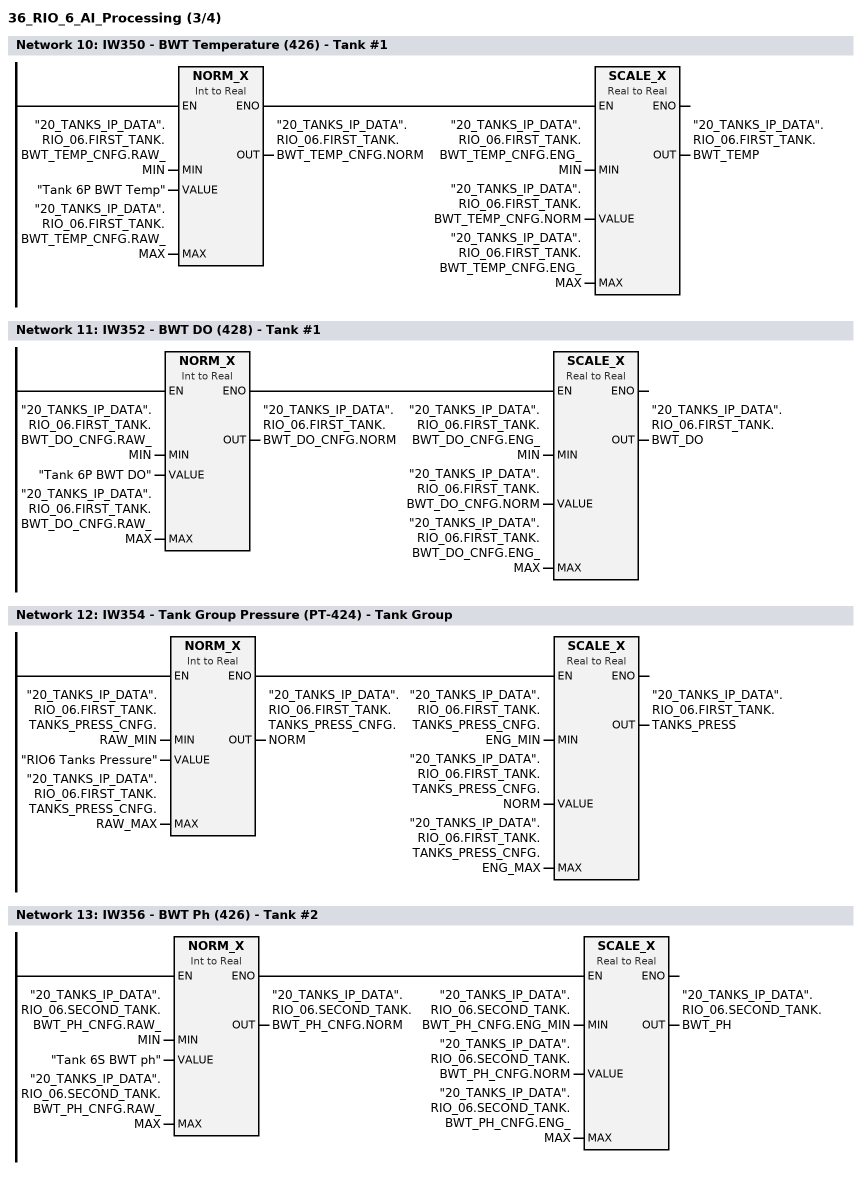
   RUNG wire#powerrail
      { S7_Templates := "[SrcType := Int, DestType := Real]" } Normalize(min := "20_TANKS_IP_DATA".RIO_06.FIRST_TANK.BWT_TEMP_CNFG.RAW_MIN, value := "Tank 6P BWT Temp", max := "20_TANKS_IP_DATA".RIO_06.FIRST_TANK.BWT_TEMP_CNFG.RAW_MAX, out => "20_TANKS_IP_DATA".RIO_06.FIRST_TANK.BWT_TEMP_CNFG.NORM)
      { S7_Templates := "[SrcType := Real, DestType := Real]" } Scale(min := "20_TANKS_IP_DATA".RIO_06.FIRST_TANK.BWT_TEMP_CNFG.ENG_MIN, value := "20_TANKS_IP_DATA".RIO_06.FIRST_TANK.BWT_TEMP_CNFG.NORM, max := "20_TANKS_IP_DATA".RIO_06.FIRST_TANK.BWT_TEMP_CNFG.ENG_MAX, out => "20_TANKS_IP_DATA".RIO_06.FIRST_TANK.BWT_TEMP)
   END_RUNG
   // the same network as SCL:
   "20_TANKS_IP_DATA".RIO_06.FIRST_TANK.BWT_TEMP_CNFG.NORM := NORM_X(MIN := "20_TANKS_IP_DATA".RIO_06.FIRST_TANK.BWT_TEMP_CNFG.RAW_MIN, VALUE := "Tank 6P BWT Temp", MAX := "20_TANKS_IP_DATA".RIO_06.FIRST_TANK.BWT_TEMP_CNFG.RAW_MAX);
   "20_TANKS_IP_DATA".RIO_06.FIRST_TANK.BWT_TEMP := SCALE_X(MIN := "20_TANKS_IP_DATA".RIO_06.FIRST_TANK.BWT_TEMP_CNFG.ENG_MIN, VALUE := "20_TANKS_IP_DATA".RIO_06.FIRST_TANK.BWT_TEMP_CNFG.NORM, MAX := "20_TANKS_IP_DATA".RIO_06.FIRST_TANK.BWT_TEMP_CNFG.ENG_MAX);
END_REGION

REGION Network 11: IW352 - BWT DO (428) - Tank #1
   RUNG wire#powerrail
      { S7_Templates := "[SrcType := Int, DestType := Real]" } Normalize(min := "20_TANKS_IP_DATA".RIO_06.FIRST_TANK.BWT_DO_CNFG.RAW_MIN, value := "Tank 6P BWT DO", max := "20_TANKS_IP_DATA".RIO_06.FIRST_TANK.BWT_DO_CNFG.RAW_MAX, out => "20_TANKS_IP_DATA".RIO_06.FIRST_TANK.BWT_DO_CNFG.NORM)
      { S7_Templates := "[SrcType := Real, DestType := Real]" } Scale(min := "20_TANKS_IP_DATA".RIO_06.FIRST_TANK.BWT_DO_CNFG.ENG_MIN, value := "20_TANKS_IP_DATA".RIO_06.FIRST_TANK.BWT_DO_CNFG.NORM, max := "20_TANKS_IP_DATA".RIO_06.FIRST_TANK.BWT_DO_CNFG.ENG_MAX, out => "20_TANKS_IP_DATA".RIO_06.FIRST_TANK.BWT_DO)
   END_RUNG
   // the same network as SCL:
   "20_TANKS_IP_DATA".RIO_06.FIRST_TANK.BWT_DO_CNFG.NORM := NORM_X(MIN := "20_TANKS_IP_DATA".RIO_06.FIRST_TANK.BWT_DO_CNFG.RAW_MIN, VALUE := "Tank 6P BWT DO", MAX := "20_TANKS_IP_DATA".RIO_06.FIRST_TANK.BWT_DO_CNFG.RAW_MAX);
   "20_TANKS_IP_DATA".RIO_06.FIRST_TANK.BWT_DO := SCALE_X(MIN := "20_TANKS_IP_DATA".RIO_06.FIRST_TANK.BWT_DO_CNFG.ENG_MIN, VALUE := "20_TANKS_IP_DATA".RIO_06.FIRST_TANK.BWT_DO_CNFG.NORM, MAX := "20_TANKS_IP_DATA".RIO_06.FIRST_TANK.BWT_DO_CNFG.ENG_MAX);
END_REGION

REGION Network 12: IW354 - Tank Group Pressure (PT-424) - Tank Group
   RUNG wire#powerrail
      { S7_Templates := "[SrcType := Int, DestType := Real]" } Normalize(min := "20_TANKS_IP_DATA".RIO_06.FIRST_TANK.TANKS_PRESS_CNFG.RAW_MIN, value := "RIO6 Tanks Pressure", max := "20_TANKS_IP_DATA".RIO_06.FIRST_TANK.TANKS_PRESS_CNFG.RAW_MAX, out => "20_TANKS_IP_DATA".RIO_06.FIRST_TANK.TANKS_PRESS_CNFG.NORM)
      { S7_Templates := "[SrcType := Real, DestType := Real]" } Scale(min := "20_TANKS_IP_DATA".RIO_06.FIRST_TANK.TANKS_PRESS_CNFG.ENG_MIN, value := "20_TANKS_IP_DATA".RIO_06.FIRST_TANK.TANKS_PRESS_CNFG.NORM, max := "20_TANKS_IP_DATA".RIO_06.FIRST_TANK.TANKS_PRESS_CNFG.ENG_MAX, out => "20_TANKS_IP_DATA".RIO_06.FIRST_TANK.TANKS_PRESS)
   END_RUNG
   // the same network as SCL:
   "20_TANKS_IP_DATA".RIO_06.FIRST_TANK.TANKS_PRESS_CNFG.NORM := NORM_X(MIN := "20_TANKS_IP_DATA".RIO_06.FIRST_TANK.TANKS_PRESS_CNFG.RAW_MIN, VALUE := "RIO6 Tanks Pressure", MAX := "20_TANKS_IP_DATA".RIO_06.FIRST_TANK.TANKS_PRESS_CNFG.RAW_MAX);
   "20_TANKS_IP_DATA".RIO_06.FIRST_TANK.TANKS_PRESS := SCALE_X(MIN := "20_TANKS_IP_DATA".RIO_06.FIRST_TANK.TANKS_PRESS_CNFG.ENG_MIN, VALUE := "20_TANKS_IP_DATA".RIO_06.FIRST_TANK.TANKS_PRESS_CNFG.NORM, MAX := "20_TANKS_IP_DATA".RIO_06.FIRST_TANK.TANKS_PRESS_CNFG.ENG_MAX);
END_REGION

REGION Network 13: IW356 - BWT Ph (426) - Tank #2
   RUNG wire#powerrail
      { S7_Templates := "[SrcType := Int, DestType := Real]" } Normalize(min := "20_TANKS_IP_DATA".RIO_06.SECOND_TANK.BWT_PH_CNFG.RAW_MIN, value := "Tank 6S BWT ph", max := "20_TANKS_IP_DATA".RIO_06.SECOND_TANK.BWT_PH_CNFG.RAW_MAX, out => "20_TANKS_IP_DATA".RIO_06.SECOND_TANK.BWT_PH_CNFG.NORM)
      { S7_Templates := "[SrcType := Real, DestType := Real]" } Scale(min := "20_TANKS_IP_DATA".RIO_06.SECOND_TANK.BWT_PH_CNFG.ENG_MIN, value := "20_TANKS_IP_DATA".RIO_06.SECOND_TANK.BWT_PH_CNFG.NORM, max := "20_TANKS_IP_DATA".RIO_06.SECOND_TANK.BWT_PH_CNFG.ENG_MAX, out => "20_TANKS_IP_DATA".RIO_06.SECOND_TANK.BWT_PH)
   END_RUNG
   // the same network as SCL:
   "20_TANKS_IP_DATA".RIO_06.SECOND_TANK.BWT_PH_CNFG.NORM := NORM_X(MIN := "20_TANKS_IP_DATA".RIO_06.SECOND_TANK.BWT_PH_CNFG.RAW_MIN, VALUE := "Tank 6S BWT ph", MAX := "20_TANKS_IP_DATA".RIO_06.SECOND_TANK.BWT_PH_CNFG.RAW_MAX);
   "20_TANKS_IP_DATA".RIO_06.SECOND_TANK.BWT_PH := SCALE_X(MIN := "20_TANKS_IP_DATA".RIO_06.SECOND_TANK.BWT_PH_CNFG.ENG_MIN, VALUE := "20_TANKS_IP_DATA".RIO_06.SECOND_TANK.BWT_PH_CNFG.NORM, MAX := "20_TANKS_IP_DATA".RIO_06.SECOND_TANK.BWT_PH_CNFG.ENG_MAX);
END_REGION

REGION Network 14: IW358 - BWT Temperature (426) - Tank #2
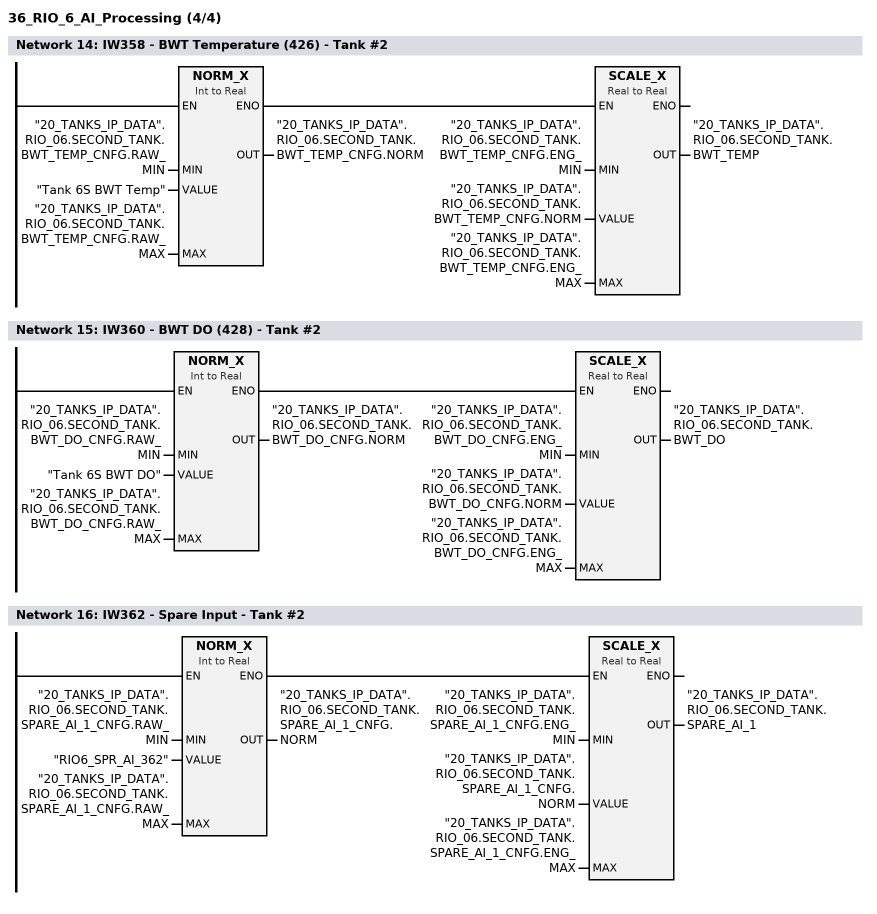
   RUNG wire#powerrail
      { S7_Templates := "[SrcType := Int, DestType := Real]" } Normalize(min := "20_TANKS_IP_DATA".RIO_06.SECOND_TANK.BWT_TEMP_CNFG.RAW_MIN, value := "Tank 6S BWT Temp", max := "20_TANKS_IP_DATA".RIO_06.SECOND_TANK.BWT_TEMP_CNFG.RAW_MAX, out => "20_TANKS_IP_DATA".RIO_06.SECOND_TANK.BWT_TEMP_CNFG.NORM)
      { S7_Templates := "[SrcType := Real, DestType := Real]" } Scale(min := "20_TANKS_IP_DATA".RIO_06.SECOND_TANK.BWT_TEMP_CNFG.ENG_MIN, value := "20_TANKS_IP_DATA".RIO_06.SECOND_TANK.BWT_TEMP_CNFG.NORM, max := "20_TANKS_IP_DATA".RIO_06.SECOND_TANK.BWT_TEMP_CNFG.ENG_MAX, out => "20_TANKS_IP_DATA".RIO_06.SECOND_TANK.BWT_TEMP)
   END_RUNG
   // the same network as SCL:
   "20_TANKS_IP_DATA".RIO_06.SECOND_TANK.BWT_TEMP_CNFG.NORM := NORM_X(MIN := "20_TANKS_IP_DATA".RIO_06.SECOND_TANK.BWT_TEMP_CNFG.RAW_MIN, VALUE := "Tank 6S BWT Temp", MAX := "20_TANKS_IP_DATA".RIO_06.SECOND_TANK.BWT_TEMP_CNFG.RAW_MAX);
   "20_TANKS_IP_DATA".RIO_06.SECOND_TANK.BWT_TEMP := SCALE_X(MIN := "20_TANKS_IP_DATA".RIO_06.SECOND_TANK.BWT_TEMP_CNFG.ENG_MIN, VALUE := "20_TANKS_IP_DATA".RIO_06.SECOND_TANK.BWT_TEMP_CNFG.NORM, MAX := "20_TANKS_IP_DATA".RIO_06.SECOND_TANK.BWT_TEMP_CNFG.ENG_MAX);
END_REGION

REGION Network 15: IW360 - BWT DO (428) - Tank #2
   RUNG wire#powerrail
      { S7_Templates := "[SrcType := Int, DestType := Real]" } Normalize(min := "20_TANKS_IP_DATA".RIO_06.SECOND_TANK.BWT_DO_CNFG.RAW_MIN, value := "Tank 6S BWT DO", max := "20_TANKS_IP_DATA".RIO_06.SECOND_TANK.BWT_DO_CNFG.RAW_MAX, out => "20_TANKS_IP_DATA".RIO_06.SECOND_TANK.BWT_DO_CNFG.NORM)
      { S7_Templates := "[SrcType := Real, DestType := Real]" } Scale(min := "20_TANKS_IP_DATA".RIO_06.SECOND_TANK.BWT_DO_CNFG.ENG_MIN, value := "20_TANKS_IP_DATA".RIO_06.SECOND_TANK.BWT_DO_CNFG.NORM, max := "20_TANKS_IP_DATA".RIO_06.SECOND_TANK.BWT_DO_CNFG.ENG_MAX, out => "20_TANKS_IP_DATA".RIO_06.SECOND_TANK.BWT_DO)
   END_RUNG
   // the same network as SCL:
   "20_TANKS_IP_DATA".RIO_06.SECOND_TANK.BWT_DO_CNFG.NORM := NORM_X(MIN := "20_TANKS_IP_DATA".RIO_06.SECOND_TANK.BWT_DO_CNFG.RAW_MIN, VALUE := "Tank 6S BWT DO", MAX := "20_TANKS_IP_DATA".RIO_06.SECOND_TANK.BWT_DO_CNFG.RAW_MAX);
   "20_TANKS_IP_DATA".RIO_06.SECOND_TANK.BWT_DO := SCALE_X(MIN := "20_TANKS_IP_DATA".RIO_06.SECOND_TANK.BWT_DO_CNFG.ENG_MIN, VALUE := "20_TANKS_IP_DATA".RIO_06.SECOND_TANK.BWT_DO_CNFG.NORM, MAX := "20_TANKS_IP_DATA".RIO_06.SECOND_TANK.BWT_DO_CNFG.ENG_MAX);
END_REGION

REGION Network 16: IW362 - Spare Input - Tank #2
   RUNG wire#powerrail
      { S7_Templates := "[SrcType := Int, DestType := Real]" } Normalize(min := "20_TANKS_IP_DATA".RIO_06.SECOND_TANK.SPARE_AI_1_CNFG.RAW_MIN, value := "RIO6_SPR_AI_362", max := "20_TANKS_IP_DATA".RIO_06.SECOND_TANK.SPARE_AI_1_CNFG.RAW_MAX, out => "20_TANKS_IP_DATA".RIO_06.SECOND_TANK.SPARE_AI_1_CNFG.NORM)
      { S7_Templates := "[SrcType := Real, DestType := Real]" } Scale(min := "20_TANKS_IP_DATA".RIO_06.SECOND_TANK.SPARE_AI_1_CNFG.ENG_MIN, value := "20_TANKS_IP_DATA".RIO_06.SECOND_TANK.SPARE_AI_1_CNFG.NORM, max := "20_TANKS_IP_DATA".RIO_06.SECOND_TANK.SPARE_AI_1_CNFG.ENG_MAX, out => "20_TANKS_IP_DATA".RIO_06.SECOND_TANK.SPARE_AI_1)
   END_RUNG
   // the same network as SCL:
   "20_TANKS_IP_DATA".RIO_06.SECOND_TANK.SPARE_AI_1_CNFG.NORM := NORM_X(MIN := "20_TANKS_IP_DATA".RIO_06.SECOND_TANK.SPARE_AI_1_CNFG.RAW_MIN, VALUE := "RIO6_SPR_AI_362", MAX := "20_TANKS_IP_DATA".RIO_06.SECOND_TANK.SPARE_AI_1_CNFG.RAW_MAX);
   "20_TANKS_IP_DATA".RIO_06.SECOND_TANK.SPARE_AI_1 := SCALE_X(MIN := "20_TANKS_IP_DATA".RIO_06.SECOND_TANK.SPARE_AI_1_CNFG.ENG_MIN, VALUE := "20_TANKS_IP_DATA".RIO_06.SECOND_TANK.SPARE_AI_1_CNFG.NORM, MAX := "20_TANKS_IP_DATA".RIO_06.SECOND_TANK.SPARE_AI_1_CNFG.ENG_MAX);
END_REGION
END_FUNCTION

FUNCTION "37_RIO_7_AI_Processing" : Void   // FC37, LAD
TITLE = Analogue Input Processing (Tank 1 = APT)
{ S7_Optimized_Access := 'TRUE' }
AUTHOR : JRS
VERSION : 0.1
// To process raw inputs prior to code use
BEGIN

REGION Network 1: IW400 - USD Flow (FIT-418) - Tank #1
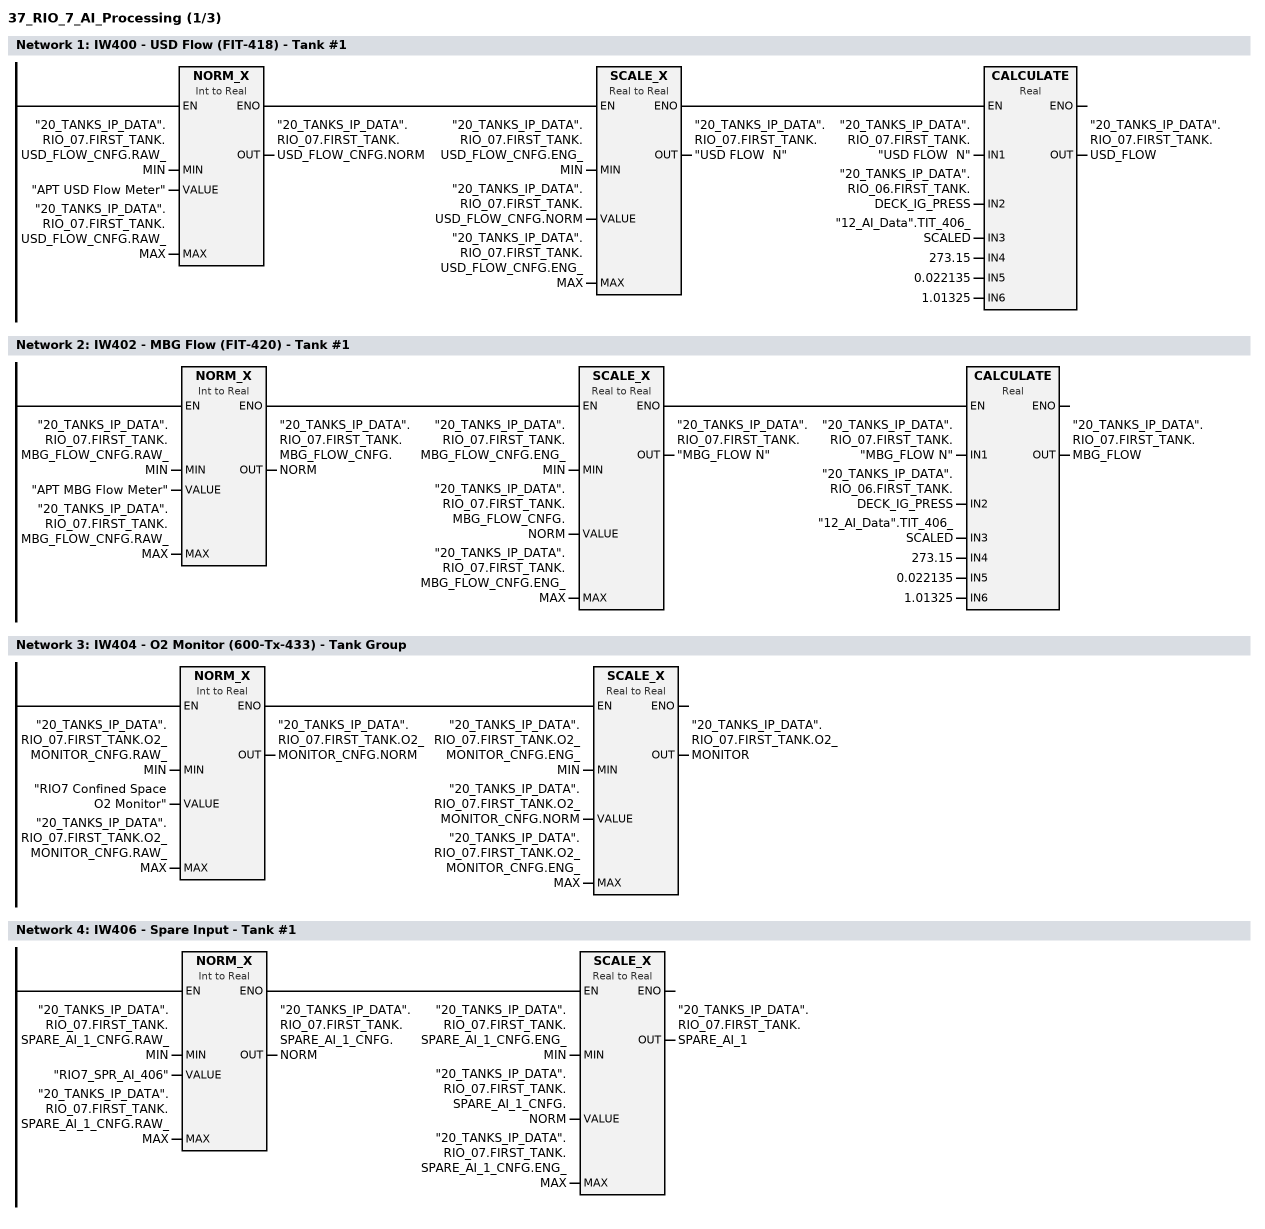
   RUNG wire#powerrail
      { S7_Templates := "[SrcType := Int, DestType := Real]" } Normalize(min := "20_TANKS_IP_DATA".RIO_07.FIRST_TANK.USD_FLOW_CNFG.RAW_MIN, value := "APT USD Flow Meter", max := "20_TANKS_IP_DATA".RIO_07.FIRST_TANK.USD_FLOW_CNFG.RAW_MAX, out => "20_TANKS_IP_DATA".RIO_07.FIRST_TANK.USD_FLOW_CNFG.NORM)
      { S7_Templates := "[SrcType := Real, DestType := Real]" } Scale(min := "20_TANKS_IP_DATA".RIO_07.FIRST_TANK.USD_FLOW_CNFG.ENG_MIN, value := "20_TANKS_IP_DATA".RIO_07.FIRST_TANK.USD_FLOW_CNFG.NORM, max := "20_TANKS_IP_DATA".RIO_07.FIRST_TANK.USD_FLOW_CNFG.ENG_MAX, out => "20_TANKS_IP_DATA".RIO_07.FIRST_TANK."USD FLOW  N")
      { S7_Templates := "SrcType := Real"; S7_Expression := "IN1*(IN2+IN6)/IN6*IN4/(IN3+IN4)" } Calculate(in1 := "20_TANKS_IP_DATA".RIO_07.FIRST_TANK."USD FLOW  N", in2 := "20_TANKS_IP_DATA".RIO_06.FIRST_TANK.DECK_IG_PRESS, in3 := "12_AI_Data".TIT_406_SCALED, in4 := 273.15, in5 := 0.022135, in6 := 1.01325, out => "20_TANKS_IP_DATA".RIO_07.FIRST_TANK.USD_FLOW)
   END_RUNG
   // the same network as SCL:
   "20_TANKS_IP_DATA".RIO_07.FIRST_TANK.USD_FLOW_CNFG.NORM := NORM_X(MIN := "20_TANKS_IP_DATA".RIO_07.FIRST_TANK.USD_FLOW_CNFG.RAW_MIN, VALUE := "APT USD Flow Meter", MAX := "20_TANKS_IP_DATA".RIO_07.FIRST_TANK.USD_FLOW_CNFG.RAW_MAX);
   "20_TANKS_IP_DATA".RIO_07.FIRST_TANK."USD FLOW  N" := SCALE_X(MIN := "20_TANKS_IP_DATA".RIO_07.FIRST_TANK.USD_FLOW_CNFG.ENG_MIN, VALUE := "20_TANKS_IP_DATA".RIO_07.FIRST_TANK.USD_FLOW_CNFG.NORM, MAX := "20_TANKS_IP_DATA".RIO_07.FIRST_TANK.USD_FLOW_CNFG.ENG_MAX);
   "20_TANKS_IP_DATA".RIO_07.FIRST_TANK.USD_FLOW := "20_TANKS_IP_DATA".RIO_07.FIRST_TANK."USD FLOW  N"*("20_TANKS_IP_DATA".RIO_06.FIRST_TANK.DECK_IG_PRESS+1.01325)/1.01325*273.15/("12_AI_Data".TIT_406_SCALED+273.15);
END_REGION

REGION Network 2: IW402 - MBG Flow (FIT-420) - Tank #1
   RUNG wire#powerrail
      { S7_Templates := "[SrcType := Int, DestType := Real]" } Normalize(min := "20_TANKS_IP_DATA".RIO_07.FIRST_TANK.MBG_FLOW_CNFG.RAW_MIN, value := "APT MBG Flow Meter", max := "20_TANKS_IP_DATA".RIO_07.FIRST_TANK.MBG_FLOW_CNFG.RAW_MAX, out => "20_TANKS_IP_DATA".RIO_07.FIRST_TANK.MBG_FLOW_CNFG.NORM)
      { S7_Templates := "[SrcType := Real, DestType := Real]" } Scale(min := "20_TANKS_IP_DATA".RIO_07.FIRST_TANK.MBG_FLOW_CNFG.ENG_MIN, value := "20_TANKS_IP_DATA".RIO_07.FIRST_TANK.MBG_FLOW_CNFG.NORM, max := "20_TANKS_IP_DATA".RIO_07.FIRST_TANK.MBG_FLOW_CNFG.ENG_MAX, out => "20_TANKS_IP_DATA".RIO_07.FIRST_TANK."MBG_FLOW N")
      { S7_Templates := "SrcType := Real"; S7_Expression := "IN1*(IN2+IN6)/IN6*IN4/(IN3+IN4)" } Calculate(in1 := "20_TANKS_IP_DATA".RIO_07.FIRST_TANK."MBG_FLOW N", in2 := "20_TANKS_IP_DATA".RIO_06.FIRST_TANK.DECK_IG_PRESS, in3 := "12_AI_Data".TIT_406_SCALED, in4 := 273.15, in5 := 0.022135, in6 := 1.01325, out => "20_TANKS_IP_DATA".RIO_07.FIRST_TANK.MBG_FLOW)
   END_RUNG
   // the same network as SCL:
   "20_TANKS_IP_DATA".RIO_07.FIRST_TANK.MBG_FLOW_CNFG.NORM := NORM_X(MIN := "20_TANKS_IP_DATA".RIO_07.FIRST_TANK.MBG_FLOW_CNFG.RAW_MIN, VALUE := "APT MBG Flow Meter", MAX := "20_TANKS_IP_DATA".RIO_07.FIRST_TANK.MBG_FLOW_CNFG.RAW_MAX);
   "20_TANKS_IP_DATA".RIO_07.FIRST_TANK."MBG_FLOW N" := SCALE_X(MIN := "20_TANKS_IP_DATA".RIO_07.FIRST_TANK.MBG_FLOW_CNFG.ENG_MIN, VALUE := "20_TANKS_IP_DATA".RIO_07.FIRST_TANK.MBG_FLOW_CNFG.NORM, MAX := "20_TANKS_IP_DATA".RIO_07.FIRST_TANK.MBG_FLOW_CNFG.ENG_MAX);
   "20_TANKS_IP_DATA".RIO_07.FIRST_TANK.MBG_FLOW := "20_TANKS_IP_DATA".RIO_07.FIRST_TANK."MBG_FLOW N"*("20_TANKS_IP_DATA".RIO_06.FIRST_TANK.DECK_IG_PRESS+1.01325)/1.01325*273.15/("12_AI_Data".TIT_406_SCALED+273.15);
END_REGION

REGION Network 3: IW404 - O2 Monitor (600-Tx-433) - Tank Group
   RUNG wire#powerrail
      { S7_Templates := "[SrcType := Int, DestType := Real]" } Normalize(min := "20_TANKS_IP_DATA".RIO_07.FIRST_TANK.O2_MONITOR_CNFG.RAW_MIN, value := "RIO7 Confined Space O2 Monitor", max := "20_TANKS_IP_DATA".RIO_07.FIRST_TANK.O2_MONITOR_CNFG.RAW_MAX, out => "20_TANKS_IP_DATA".RIO_07.FIRST_TANK.O2_MONITOR_CNFG.NORM)
      { S7_Templates := "[SrcType := Real, DestType := Real]" } Scale(min := "20_TANKS_IP_DATA".RIO_07.FIRST_TANK.O2_MONITOR_CNFG.ENG_MIN, value := "20_TANKS_IP_DATA".RIO_07.FIRST_TANK.O2_MONITOR_CNFG.NORM, max := "20_TANKS_IP_DATA".RIO_07.FIRST_TANK.O2_MONITOR_CNFG.ENG_MAX, out => "20_TANKS_IP_DATA".RIO_07.FIRST_TANK.O2_MONITOR)
   END_RUNG
   // the same network as SCL:
   "20_TANKS_IP_DATA".RIO_07.FIRST_TANK.O2_MONITOR_CNFG.NORM := NORM_X(MIN := "20_TANKS_IP_DATA".RIO_07.FIRST_TANK.O2_MONITOR_CNFG.RAW_MIN, VALUE := "RIO7 Confined Space O2 Monitor", MAX := "20_TANKS_IP_DATA".RIO_07.FIRST_TANK.O2_MONITOR_CNFG.RAW_MAX);
   "20_TANKS_IP_DATA".RIO_07.FIRST_TANK.O2_MONITOR := SCALE_X(MIN := "20_TANKS_IP_DATA".RIO_07.FIRST_TANK.O2_MONITOR_CNFG.ENG_MIN, VALUE := "20_TANKS_IP_DATA".RIO_07.FIRST_TANK.O2_MONITOR_CNFG.NORM, MAX := "20_TANKS_IP_DATA".RIO_07.FIRST_TANK.O2_MONITOR_CNFG.ENG_MAX);
END_REGION

REGION Network 4: IW406 - Spare Input - Tank #1
   RUNG wire#powerrail
      { S7_Templates := "[SrcType := Int, DestType := Real]" } Normalize(min := "20_TANKS_IP_DATA".RIO_07.FIRST_TANK.SPARE_AI_1_CNFG.RAW_MIN, value := "RIO7_SPR_AI_406", max := "20_TANKS_IP_DATA".RIO_07.FIRST_TANK.SPARE_AI_1_CNFG.RAW_MAX, out => "20_TANKS_IP_DATA".RIO_07.FIRST_TANK.SPARE_AI_1_CNFG.NORM)
      { S7_Templates := "[SrcType := Real, DestType := Real]" } Scale(min := "20_TANKS_IP_DATA".RIO_07.FIRST_TANK.SPARE_AI_1_CNFG.ENG_MIN, value := "20_TANKS_IP_DATA".RIO_07.FIRST_TANK.SPARE_AI_1_CNFG.NORM, max := "20_TANKS_IP_DATA".RIO_07.FIRST_TANK.SPARE_AI_1_CNFG.ENG_MAX, out => "20_TANKS_IP_DATA".RIO_07.FIRST_TANK.SPARE_AI_1)
   END_RUNG
   // the same network as SCL:
   "20_TANKS_IP_DATA".RIO_07.FIRST_TANK.SPARE_AI_1_CNFG.NORM := NORM_X(MIN := "20_TANKS_IP_DATA".RIO_07.FIRST_TANK.SPARE_AI_1_CNFG.RAW_MIN, VALUE := "RIO7_SPR_AI_406", MAX := "20_TANKS_IP_DATA".RIO_07.FIRST_TANK.SPARE_AI_1_CNFG.RAW_MAX);
   "20_TANKS_IP_DATA".RIO_07.FIRST_TANK.SPARE_AI_1 := SCALE_X(MIN := "20_TANKS_IP_DATA".RIO_07.FIRST_TANK.SPARE_AI_1_CNFG.ENG_MIN, VALUE := "20_TANKS_IP_DATA".RIO_07.FIRST_TANK.SPARE_AI_1_CNFG.NORM, MAX := "20_TANKS_IP_DATA".RIO_07.FIRST_TANK.SPARE_AI_1_CNFG.ENG_MAX);
END_REGION

REGION Network 5: IW408 - Deck Main IG Pressure (PT-415) - Tank Group
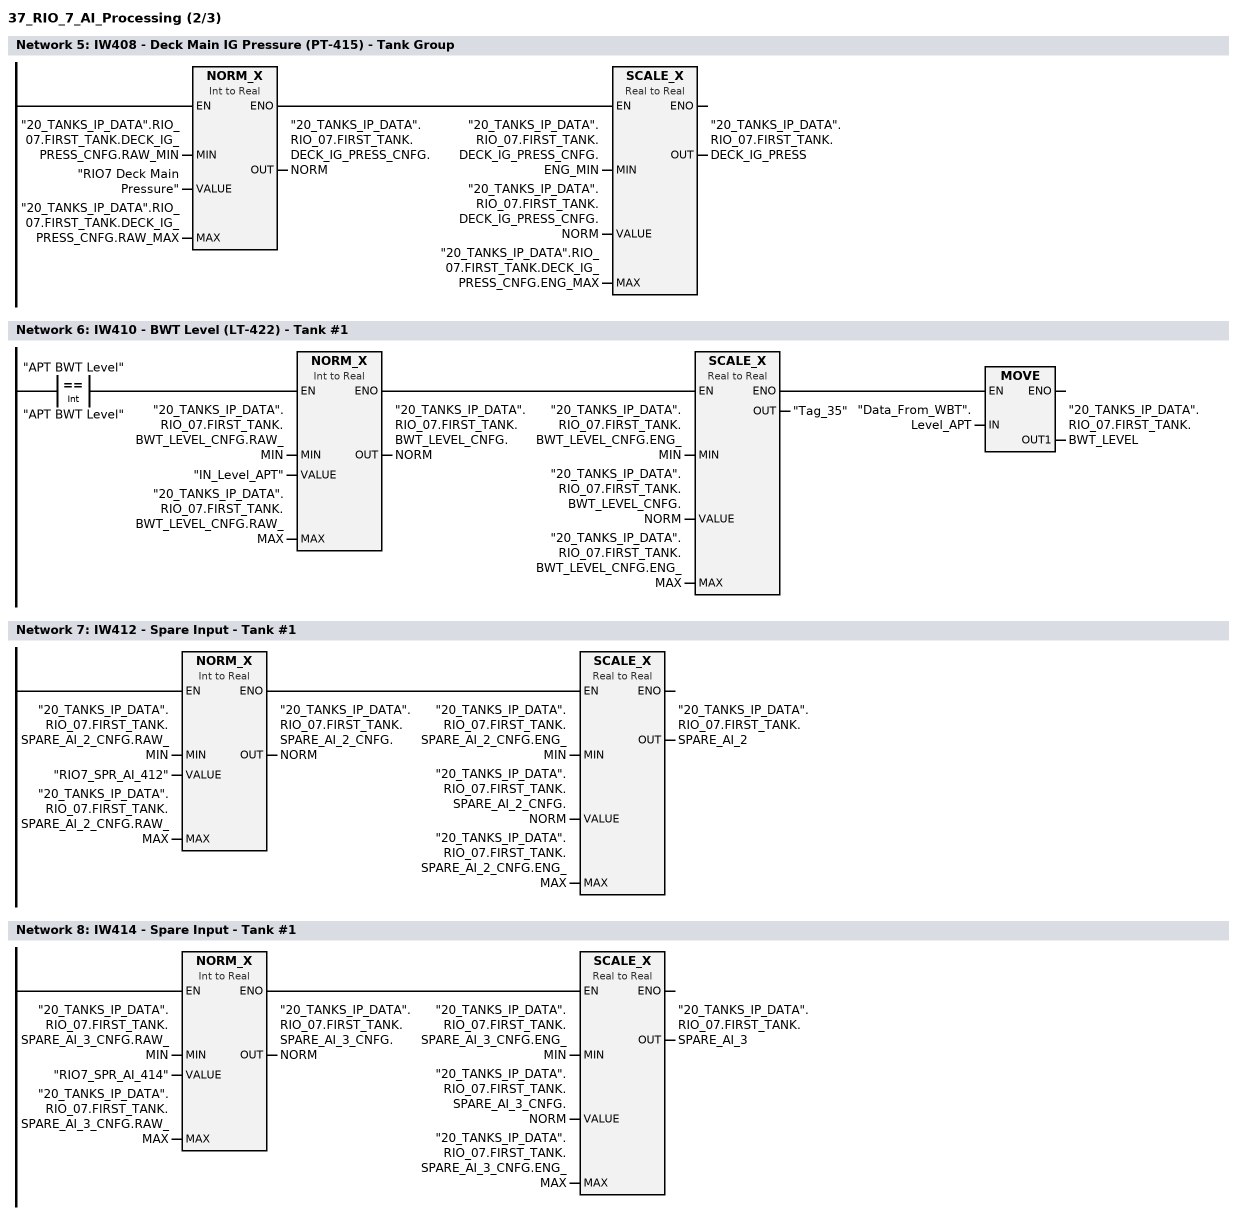
   RUNG wire#powerrail
      { S7_Templates := "[SrcType := Int, DestType := Real]" } Normalize(min := "20_TANKS_IP_DATA".RIO_07.FIRST_TANK.DECK_IG_PRESS_CNFG.RAW_MIN, value := "RIO7 Deck Main Pressure", max := "20_TANKS_IP_DATA".RIO_07.FIRST_TANK.DECK_IG_PRESS_CNFG.RAW_MAX, out => "20_TANKS_IP_DATA".RIO_07.FIRST_TANK.DECK_IG_PRESS_CNFG.NORM)
      { S7_Templates := "[SrcType := Real, DestType := Real]" } Scale(min := "20_TANKS_IP_DATA".RIO_07.FIRST_TANK.DECK_IG_PRESS_CNFG.ENG_MIN, value := "20_TANKS_IP_DATA".RIO_07.FIRST_TANK.DECK_IG_PRESS_CNFG.NORM, max := "20_TANKS_IP_DATA".RIO_07.FIRST_TANK.DECK_IG_PRESS_CNFG.ENG_MAX, out => "20_TANKS_IP_DATA".RIO_07.FIRST_TANK.DECK_IG_PRESS)
   END_RUNG
   // the same network as SCL:
   "20_TANKS_IP_DATA".RIO_07.FIRST_TANK.DECK_IG_PRESS_CNFG.NORM := NORM_X(MIN := "20_TANKS_IP_DATA".RIO_07.FIRST_TANK.DECK_IG_PRESS_CNFG.RAW_MIN, VALUE := "RIO7 Deck Main Pressure", MAX := "20_TANKS_IP_DATA".RIO_07.FIRST_TANK.DECK_IG_PRESS_CNFG.RAW_MAX);
   "20_TANKS_IP_DATA".RIO_07.FIRST_TANK.DECK_IG_PRESS := SCALE_X(MIN := "20_TANKS_IP_DATA".RIO_07.FIRST_TANK.DECK_IG_PRESS_CNFG.ENG_MIN, VALUE := "20_TANKS_IP_DATA".RIO_07.FIRST_TANK.DECK_IG_PRESS_CNFG.NORM, MAX := "20_TANKS_IP_DATA".RIO_07.FIRST_TANK.DECK_IG_PRESS_CNFG.ENG_MAX);
END_REGION

REGION Network 6: IW410 - BWT Level (LT-422) - Tank #1
   RUNG wire#powerrail
      { S7_Templates := "SrcType := Int" } EQ_Contact(in1 := "APT BWT Level", in2 := "APT BWT Level")
      { S7_Templates := "[SrcType := Int, DestType := Real]" } Normalize(min := "20_TANKS_IP_DATA".RIO_07.FIRST_TANK.BWT_LEVEL_CNFG.RAW_MIN, value := "IN_Level_APT", max := "20_TANKS_IP_DATA".RIO_07.FIRST_TANK.BWT_LEVEL_CNFG.RAW_MAX, out => "20_TANKS_IP_DATA".RIO_07.FIRST_TANK.BWT_LEVEL_CNFG.NORM)
      { S7_Templates := "[SrcType := Real, DestType := Real]" } Scale(min := "20_TANKS_IP_DATA".RIO_07.FIRST_TANK.BWT_LEVEL_CNFG.ENG_MIN, value := "20_TANKS_IP_DATA".RIO_07.FIRST_TANK.BWT_LEVEL_CNFG.NORM, max := "20_TANKS_IP_DATA".RIO_07.FIRST_TANK.BWT_LEVEL_CNFG.ENG_MAX, out => "Tag_35")
      Move(in := "Data_From_WBT".Level_APT, out1 => "20_TANKS_IP_DATA".RIO_07.FIRST_TANK.BWT_LEVEL)
   END_RUNG
   // the same network as SCL:
   IF "APT BWT Level" = "APT BWT Level" THEN
       "20_TANKS_IP_DATA".RIO_07.FIRST_TANK.BWT_LEVEL_CNFG.NORM := NORM_X(MIN := "20_TANKS_IP_DATA".RIO_07.FIRST_TANK.BWT_LEVEL_CNFG.RAW_MIN, VALUE := "IN_Level_APT", MAX := "20_TANKS_IP_DATA".RIO_07.FIRST_TANK.BWT_LEVEL_CNFG.RAW_MAX);
       "Tag_35" := SCALE_X(MIN := "20_TANKS_IP_DATA".RIO_07.FIRST_TANK.BWT_LEVEL_CNFG.ENG_MIN, VALUE := "20_TANKS_IP_DATA".RIO_07.FIRST_TANK.BWT_LEVEL_CNFG.NORM, MAX := "20_TANKS_IP_DATA".RIO_07.FIRST_TANK.BWT_LEVEL_CNFG.ENG_MAX);
       "20_TANKS_IP_DATA".RIO_07.FIRST_TANK.BWT_LEVEL := "Data_From_WBT".Level_APT;
   END_IF;
END_REGION

REGION Network 7: IW412 - Spare Input - Tank #1
   RUNG wire#powerrail
      { S7_Templates := "[SrcType := Int, DestType := Real]" } Normalize(min := "20_TANKS_IP_DATA".RIO_07.FIRST_TANK.SPARE_AI_2_CNFG.RAW_MIN, value := "RIO7_SPR_AI_412", max := "20_TANKS_IP_DATA".RIO_07.FIRST_TANK.SPARE_AI_2_CNFG.RAW_MAX, out => "20_TANKS_IP_DATA".RIO_07.FIRST_TANK.SPARE_AI_2_CNFG.NORM)
      { S7_Templates := "[SrcType := Real, DestType := Real]" } Scale(min := "20_TANKS_IP_DATA".RIO_07.FIRST_TANK.SPARE_AI_2_CNFG.ENG_MIN, value := "20_TANKS_IP_DATA".RIO_07.FIRST_TANK.SPARE_AI_2_CNFG.NORM, max := "20_TANKS_IP_DATA".RIO_07.FIRST_TANK.SPARE_AI_2_CNFG.ENG_MAX, out => "20_TANKS_IP_DATA".RIO_07.FIRST_TANK.SPARE_AI_2)
   END_RUNG
   // the same network as SCL:
   "20_TANKS_IP_DATA".RIO_07.FIRST_TANK.SPARE_AI_2_CNFG.NORM := NORM_X(MIN := "20_TANKS_IP_DATA".RIO_07.FIRST_TANK.SPARE_AI_2_CNFG.RAW_MIN, VALUE := "RIO7_SPR_AI_412", MAX := "20_TANKS_IP_DATA".RIO_07.FIRST_TANK.SPARE_AI_2_CNFG.RAW_MAX);
   "20_TANKS_IP_DATA".RIO_07.FIRST_TANK.SPARE_AI_2 := SCALE_X(MIN := "20_TANKS_IP_DATA".RIO_07.FIRST_TANK.SPARE_AI_2_CNFG.ENG_MIN, VALUE := "20_TANKS_IP_DATA".RIO_07.FIRST_TANK.SPARE_AI_2_CNFG.NORM, MAX := "20_TANKS_IP_DATA".RIO_07.FIRST_TANK.SPARE_AI_2_CNFG.ENG_MAX);
END_REGION

REGION Network 8: IW414 - Spare Input - Tank #1
   RUNG wire#powerrail
      { S7_Templates := "[SrcType := Int, DestType := Real]" } Normalize(min := "20_TANKS_IP_DATA".RIO_07.FIRST_TANK.SPARE_AI_3_CNFG.RAW_MIN, value := "RIO7_SPR_AI_414", max := "20_TANKS_IP_DATA".RIO_07.FIRST_TANK.SPARE_AI_3_CNFG.RAW_MAX, out => "20_TANKS_IP_DATA".RIO_07.FIRST_TANK.SPARE_AI_3_CNFG.NORM)
      { S7_Templates := "[SrcType := Real, DestType := Real]" } Scale(min := "20_TANKS_IP_DATA".RIO_07.FIRST_TANK.SPARE_AI_3_CNFG.ENG_MIN, value := "20_TANKS_IP_DATA".RIO_07.FIRST_TANK.SPARE_AI_3_CNFG.NORM, max := "20_TANKS_IP_DATA".RIO_07.FIRST_TANK.SPARE_AI_3_CNFG.ENG_MAX, out => "20_TANKS_IP_DATA".RIO_07.FIRST_TANK.SPARE_AI_3)
   END_RUNG
   // the same network as SCL:
   "20_TANKS_IP_DATA".RIO_07.FIRST_TANK.SPARE_AI_3_CNFG.NORM := NORM_X(MIN := "20_TANKS_IP_DATA".RIO_07.FIRST_TANK.SPARE_AI_3_CNFG.RAW_MIN, VALUE := "RIO7_SPR_AI_414", MAX := "20_TANKS_IP_DATA".RIO_07.FIRST_TANK.SPARE_AI_3_CNFG.RAW_MAX);
   "20_TANKS_IP_DATA".RIO_07.FIRST_TANK.SPARE_AI_3 := SCALE_X(MIN := "20_TANKS_IP_DATA".RIO_07.FIRST_TANK.SPARE_AI_3_CNFG.ENG_MIN, VALUE := "20_TANKS_IP_DATA".RIO_07.FIRST_TANK.SPARE_AI_3_CNFG.NORM, MAX := "20_TANKS_IP_DATA".RIO_07.FIRST_TANK.SPARE_AI_3_CNFG.ENG_MAX);
END_REGION

REGION Network 9: IW416 - BWT Ph (426) - Tank #1
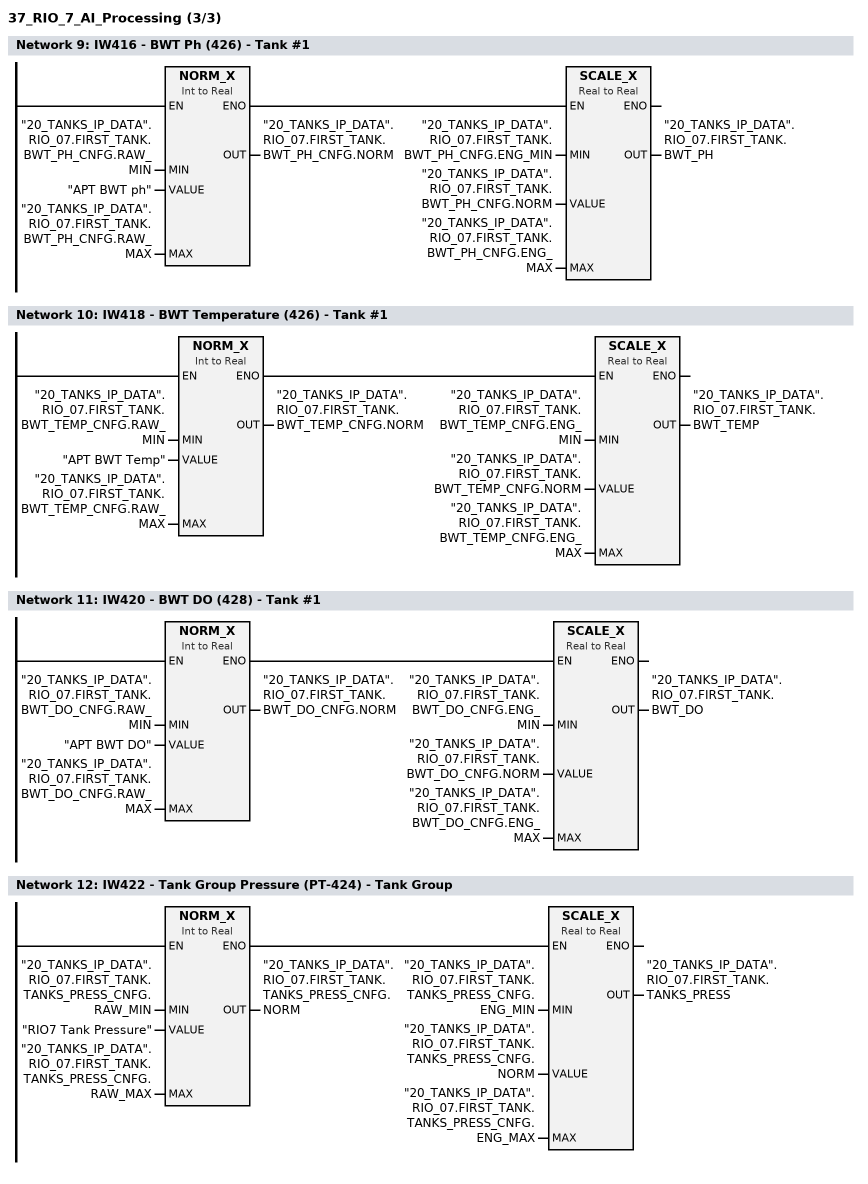
   RUNG wire#powerrail
      { S7_Templates := "[SrcType := Int, DestType := Real]" } Normalize(min := "20_TANKS_IP_DATA".RIO_07.FIRST_TANK.BWT_PH_CNFG.RAW_MIN, value := "APT BWT ph", max := "20_TANKS_IP_DATA".RIO_07.FIRST_TANK.BWT_PH_CNFG.RAW_MAX, out => "20_TANKS_IP_DATA".RIO_07.FIRST_TANK.BWT_PH_CNFG.NORM)
      { S7_Templates := "[SrcType := Real, DestType := Real]" } Scale(min := "20_TANKS_IP_DATA".RIO_07.FIRST_TANK.BWT_PH_CNFG.ENG_MIN, value := "20_TANKS_IP_DATA".RIO_07.FIRST_TANK.BWT_PH_CNFG.NORM, max := "20_TANKS_IP_DATA".RIO_07.FIRST_TANK.BWT_PH_CNFG.ENG_MAX, out => "20_TANKS_IP_DATA".RIO_07.FIRST_TANK.BWT_PH)
   END_RUNG
   // the same network as SCL:
   "20_TANKS_IP_DATA".RIO_07.FIRST_TANK.BWT_PH_CNFG.NORM := NORM_X(MIN := "20_TANKS_IP_DATA".RIO_07.FIRST_TANK.BWT_PH_CNFG.RAW_MIN, VALUE := "APT BWT ph", MAX := "20_TANKS_IP_DATA".RIO_07.FIRST_TANK.BWT_PH_CNFG.RAW_MAX);
   "20_TANKS_IP_DATA".RIO_07.FIRST_TANK.BWT_PH := SCALE_X(MIN := "20_TANKS_IP_DATA".RIO_07.FIRST_TANK.BWT_PH_CNFG.ENG_MIN, VALUE := "20_TANKS_IP_DATA".RIO_07.FIRST_TANK.BWT_PH_CNFG.NORM, MAX := "20_TANKS_IP_DATA".RIO_07.FIRST_TANK.BWT_PH_CNFG.ENG_MAX);
END_REGION

REGION Network 10: IW418 - BWT Temperature (426) - Tank #1
   RUNG wire#powerrail
      { S7_Templates := "[SrcType := Int, DestType := Real]" } Normalize(min := "20_TANKS_IP_DATA".RIO_07.FIRST_TANK.BWT_TEMP_CNFG.RAW_MIN, value := "APT BWT Temp", max := "20_TANKS_IP_DATA".RIO_07.FIRST_TANK.BWT_TEMP_CNFG.RAW_MAX, out => "20_TANKS_IP_DATA".RIO_07.FIRST_TANK.BWT_TEMP_CNFG.NORM)
      { S7_Templates := "[SrcType := Real, DestType := Real]" } Scale(min := "20_TANKS_IP_DATA".RIO_07.FIRST_TANK.BWT_TEMP_CNFG.ENG_MIN, value := "20_TANKS_IP_DATA".RIO_07.FIRST_TANK.BWT_TEMP_CNFG.NORM, max := "20_TANKS_IP_DATA".RIO_07.FIRST_TANK.BWT_TEMP_CNFG.ENG_MAX, out => "20_TANKS_IP_DATA".RIO_07.FIRST_TANK.BWT_TEMP)
   END_RUNG
   // the same network as SCL:
   "20_TANKS_IP_DATA".RIO_07.FIRST_TANK.BWT_TEMP_CNFG.NORM := NORM_X(MIN := "20_TANKS_IP_DATA".RIO_07.FIRST_TANK.BWT_TEMP_CNFG.RAW_MIN, VALUE := "APT BWT Temp", MAX := "20_TANKS_IP_DATA".RIO_07.FIRST_TANK.BWT_TEMP_CNFG.RAW_MAX);
   "20_TANKS_IP_DATA".RIO_07.FIRST_TANK.BWT_TEMP := SCALE_X(MIN := "20_TANKS_IP_DATA".RIO_07.FIRST_TANK.BWT_TEMP_CNFG.ENG_MIN, VALUE := "20_TANKS_IP_DATA".RIO_07.FIRST_TANK.BWT_TEMP_CNFG.NORM, MAX := "20_TANKS_IP_DATA".RIO_07.FIRST_TANK.BWT_TEMP_CNFG.ENG_MAX);
END_REGION

REGION Network 11: IW420 - BWT DO (428) - Tank #1
   RUNG wire#powerrail
      { S7_Templates := "[SrcType := Int, DestType := Real]" } Normalize(min := "20_TANKS_IP_DATA".RIO_07.FIRST_TANK.BWT_DO_CNFG.RAW_MIN, value := "APT BWT DO", max := "20_TANKS_IP_DATA".RIO_07.FIRST_TANK.BWT_DO_CNFG.RAW_MAX, out => "20_TANKS_IP_DATA".RIO_07.FIRST_TANK.BWT_DO_CNFG.NORM)
      { S7_Templates := "[SrcType := Real, DestType := Real]" } Scale(min := "20_TANKS_IP_DATA".RIO_07.FIRST_TANK.BWT_DO_CNFG.ENG_MIN, value := "20_TANKS_IP_DATA".RIO_07.FIRST_TANK.BWT_DO_CNFG.NORM, max := "20_TANKS_IP_DATA".RIO_07.FIRST_TANK.BWT_DO_CNFG.ENG_MAX, out => "20_TANKS_IP_DATA".RIO_07.FIRST_TANK.BWT_DO)
   END_RUNG
   // the same network as SCL:
   "20_TANKS_IP_DATA".RIO_07.FIRST_TANK.BWT_DO_CNFG.NORM := NORM_X(MIN := "20_TANKS_IP_DATA".RIO_07.FIRST_TANK.BWT_DO_CNFG.RAW_MIN, VALUE := "APT BWT DO", MAX := "20_TANKS_IP_DATA".RIO_07.FIRST_TANK.BWT_DO_CNFG.RAW_MAX);
   "20_TANKS_IP_DATA".RIO_07.FIRST_TANK.BWT_DO := SCALE_X(MIN := "20_TANKS_IP_DATA".RIO_07.FIRST_TANK.BWT_DO_CNFG.ENG_MIN, VALUE := "20_TANKS_IP_DATA".RIO_07.FIRST_TANK.BWT_DO_CNFG.NORM, MAX := "20_TANKS_IP_DATA".RIO_07.FIRST_TANK.BWT_DO_CNFG.ENG_MAX);
END_REGION

